(* Logix 5000 project; controller FV vendor 1 type 14 code 217 rev 31.11; software revision 31.00; part 61 of 63 *)
(* tags used below, declared in another part *)
   CWD : CHECKWORD_FLAGS;
   FV_N88 : INT[255];   // YSP COMMS Data transferred to/ from yeast press PLC
   One_Second_One_Scan : ALIAS FOR One_Second_1_scan;
   YP_B103 : INT[15];   // Original N File From SLC, No Description Available
   YP_BLUNG_OV : PlantItem;   // BLUNG_OV
   YP_BLUNG_OV_RawInput : ALIAS FOR RIO_Rack_3:2:I.Data.1;   // YP_BLUNG_OV
   YP_CONV_STOP : PlantItem;   // CONV_STOP
   YP_CONV_STOP_RawInput : ALIAS FOR RIO_Rack_3:2:I.Data.7;   // YP_CONV_STOP
   YP_INP1 : PlantItem;   // INP1
   YP_INP10 : PlantItem;   // INP10
   YP_INP10_RawInput : ALIAS FOR RIO_Rack_3:2:I.Data.14;   // YP_INP10
   YP_INP11 : PlantItem;   // INP11
   YP_INP11_RawInput : ALIAS FOR RIO_Rack_3:2:I.Data.15;   // YP_INP11
   YP_INP1_RawInput : ALIAS FOR RIO_Rack_3:2:I.Data.2;   // YP_INP1
   YP_INP2 : PlantItem;   // INP2
   YP_INP2_RawInput : ALIAS FOR RIO_Rack_3:2:I.Data.3;   // YP_INP2
   YP_INP3 : PlantItem;   // INP3
   YP_INP3_RawInput : ALIAS FOR RIO_Rack_3:2:I.Data.4;   // YP_INP3
   YP_INP4 : PlantItem;   // INP4
   YP_INP4_RawInput : ALIAS FOR RIO_Rack_3:2:I.Data.8;   // YP_INP4
   YP_INP5 : PlantItem;   // INP5
   YP_INP5_RawInput : ALIAS FOR RIO_Rack_3:2:I.Data.9;   // YP_INP5
   YP_INP6 : PlantItem;   // INP6
   YP_INP6_RawInput : ALIAS FOR RIO_Rack_3:2:I.Data.10;   // YP_INP6
   YP_INP7 : PlantItem;   // INP7
   YP_INP7_RawInput : ALIAS FOR RIO_Rack_3:2:I.Data.11;   // YP_INP7
   YP_INP8 : PlantItem;   // INP8
   YP_INP8_RawInput : ALIAS FOR RIO_Rack_3:2:I.Data.12;   // YP_INP8
   YP_INP9 : PlantItem;   // INP9
   YP_INP9_RawInput : ALIAS FOR RIO_Rack_3:2:I.Data.13;   // YP_INP9
   YP_N10 : INT[105];   // COMMS BLOC comms block to fv pl c
   YP_N40 : INT[9];   // Original N File From SLC, No Description Available
   YP_N55 : INT[244];   // Original N File From SLC, No Description Available
   YP_N7 : INT[56];   // INTEGER
   YP_PILZ_OK : PlantItem;   // PILZ_OK
   YP_PILZ_OK_RawInput : ALIAS FOR RIO_Rack_3:2:I.Data.0;   // YP_PILZ_OK
   YP_PRESS_CL : PlantItem;   // PRESS_CL
   YP_PRESS_CL_RawInput : ALIAS FOR RIO_Rack_3:2:I.Data.5;   // YP_PRESS_CL
   YP_PRESS_OP : PlantItem;   // PRESS_OP
   YP_PRESS_OP_RawInput : ALIAS FOR RIO_Rack_3:2:I.Data.6;   // YP_PRESS_OP
   YP_T21 : TIMER[30];
   YP_YST1_HL : PlantItem;   // YST1_HL
   YP_YST1_HL_RawInput : ALIAS FOR RIO_Rack_3:1:I.Data.1;   // YP_YST1_HL
   YP_YST2_HL : PlantItem;   // YST2_HL
   YP_YST2_HL_RawInput : ALIAS FOR RIO_Rack_3:1:I.Data.3;   // YP_YST2_HL
(* YP_Common, continued *)

ROUTINE YP_BLUNGER_14   (* ladder *)
   0: XIO(YP_N40[2].0)XIO(YP_N40[2].1)OTL(YP_N40[2].0);
   1: XIC(YP_N40[2].1)XIO(YP_B103[3].0)[GRT(YP_T21[1].ACC,YP_N55[30]) ,XIC(YP_B103[3].1) ][OTU(YP_N40[2].1) ,OTL(YP_N40[2].0) ];
   2: XIC(YP_N40[2].0)XIC(YP_B103[3].0)[OTU(YP_N40[2].0) ,OTL(YP_N40[2].1) ];
   3: EQU(YP_N55[31],0)MOV(YP_N55[32],YP_N55[30]);
   4: EQU(YP_N55[31],1)MOV(YP_N55[33],YP_N55[30]);
   5: EQU(YP_N55[31],2)MOV(YP_N55[34],YP_N55[30]);
   6: XIC(YP_N40[2].1)TON(YP_T21[1],?,?);
   7: XIO(YP_N40[3].0)XIO(YP_N40[3].1)OTL(YP_N40[3].0);
   8: XIC(YP_N40[3].1)[GRT(YP_T21[2].ACC,YP_N55[40]) ,XIC(YP_B103[3].3) ,XIC(YP_N7[38].0) ,XIC(YP_N7[38].1) ][OTU(YP_N40[3].1) ,OTL(YP_N40[3].0) ];
   9: XIC(YP_N40[3].0)XIC(YP_B103[3].2)[OTU(YP_N40[3].0) ,OTL(YP_N40[3].1) ];
   10: EQU(YP_N55[41],0)MOV(YP_N55[42],YP_N55[40]);
   11: EQU(YP_N55[41],1)MOV(YP_N55[43],YP_N55[40]);
   12: EQU(YP_N55[41],2)MOV(YP_N55[44],YP_N55[40]);
   13: XIC(YP_N40[3].1)TON(YP_T21[2],?,?);
   14: XIC(YP_N40[3].1)XIC(YP_N7[40].0)EQU(YP_N7[39],1)OTL(YP_N7[38].0);
   15: XIC(YP_N40[3].1)XIC(YP_N7[40].1)EQU(YP_N7[39],2)OTL(YP_N7[38].1);
   16: XIC(YP_N40[3].1)EQU(YP_N7[39],99)OTE(YP_N7[38].2);
END_ROUTINE

ROUTINE YP_COMMS_4   (* ladder *)
   0: XIO(YP_T21[3].DN)TON(YP_T21[3],?,?);
   1: XIC(YP_T21[3].DN)COP(FV_N88[0],YP_N10[10],2);
   2: EQU(YP_N10[11],99)MOV(99,YP_N7[39]);
   3: EQU(YP_N10[11],1)MOV(1,YP_N7[39]);
   4: EQU(YP_N10[11],2)MOV(2,YP_N7[39]);
   5: XIC(YP_N7[38].0)OTE(YP_N10[1].0);
   6: XIC(YP_N7[38].1)OTE(YP_N10[1].1);
   7: XIC(YP_N10[10].0)OTE(YP_N10[0].0);
END_ROUTINE

ROUTINE YP_Digital_Inputs   (* ladder *)
   0: [XIC(S:FS) OTU(YP_YST1_HL.CW.[CWD.MANUAL]) ,[XIC(YP_YST1_HL_RawInput) XIO(YP_YST1_HL.CW.[CWD.MANUAL]) ,XIC(YP_YST1_HL.CW.[CWD.MANDRV]) XIC(YP_YST1_HL.CW.[CWD.MANUAL]) ] OTE(YP_YST1_HL.CW.[CWD.INPUTSTATUS]) ,XIC(One_Second_One_Scan) [XIC(YP_YST1_HL.CW.[CWD.INPUTSTATUS]) XIO(YP_YST1_HL.CW.[CWD.INPUTSTATUSDEBOUNCED]) ,XIO(YP_YST1_HL.CW.[CWD.INPUTSTATUS]) XIC(YP_YST1_HL.CW.[CWD.INPUTSTATUSDEBOUNCED]) ] ADD(1,YP_YST1_HL.DebounceTimer,YP_YST1_HL.DebounceTimer) ,[XIC(YP_YST1_HL.CW.[CWD.INPUTSTATUS]) XIC(YP_YST1_HL.CW.[CWD.INPUTSTATUSDEBOUNCED]) ,XIO(YP_YST1_HL.CW.[CWD.INPUTSTATUS]) XIO(YP_YST1_HL.CW.[CWD.INPUTSTATUSDEBOUNCED]) ] CLR(YP_YST1_HL.DebounceTimer) ,GEQ(YP_YST1_HL.DebounceTimer,YP_YST1_HL.DebounceTime) XIC(YP_YST1_HL.CW.[CWD.INPUTSTATUS]) [OTL(YP_YST1_HL.CW.[CWD.INPUTSTATUSDEBOUNCED]) ,CLR(YP_YST1_HL.DebounceTimer) ] ,GEQ(YP_YST1_HL.DebounceTimer,YP_YST1_HL.DebounceTime) XIO(YP_YST1_HL.CW.[CWD.INPUTSTATUS]) [OTU(YP_YST1_HL.CW.[CWD.INPUTSTATUSDEBOUNCED]) ,CLR(YP_YST1_HL.DebounceTimer) ] ];
   1: [XIC(S:FS) OTU(YP_YST2_HL.CW.[CWD.MANUAL]) ,[XIC(YP_YST2_HL_RawInput) XIO(YP_YST2_HL.CW.[CWD.MANUAL]) ,XIC(YP_YST2_HL.CW.[CWD.MANDRV]) XIC(YP_YST2_HL.CW.[CWD.MANUAL]) ] OTE(YP_YST2_HL.CW.[CWD.INPUTSTATUS]) ,XIC(One_Second_One_Scan) [XIC(YP_YST2_HL.CW.[CWD.INPUTSTATUS]) XIO(YP_YST2_HL.CW.[CWD.INPUTSTATUSDEBOUNCED]) ,XIO(YP_YST2_HL.CW.[CWD.INPUTSTATUS]) XIC(YP_YST2_HL.CW.[CWD.INPUTSTATUSDEBOUNCED]) ] ADD(1,YP_YST2_HL.DebounceTimer,YP_YST2_HL.DebounceTimer) ,[XIC(YP_YST2_HL.CW.[CWD.INPUTSTATUS]) XIC(YP_YST2_HL.CW.[CWD.INPUTSTATUSDEBOUNCED]) ,XIO(YP_YST2_HL.CW.[CWD.INPUTSTATUS]) XIO(YP_YST2_HL.CW.[CWD.INPUTSTATUSDEBOUNCED]) ] CLR(YP_YST2_HL.DebounceTimer) ,GEQ(YP_YST2_HL.DebounceTimer,YP_YST2_HL.DebounceTime) XIC(YP_YST2_HL.CW.[CWD.INPUTSTATUS]) [OTL(YP_YST2_HL.CW.[CWD.INPUTSTATUSDEBOUNCED]) ,CLR(YP_YST2_HL.DebounceTimer) ] ,GEQ(YP_YST2_HL.DebounceTimer,YP_YST2_HL.DebounceTime) XIO(YP_YST2_HL.CW.[CWD.INPUTSTATUS]) [OTU(YP_YST2_HL.CW.[CWD.INPUTSTATUSDEBOUNCED]) ,CLR(YP_YST2_HL.DebounceTimer) ] ];
   2: [XIC(S:FS) OTU(YP_PILZ_OK.CW.[CWD.MANUAL]) ,[XIC(YP_PILZ_OK_RawInput) XIO(YP_PILZ_OK.CW.[CWD.MANUAL]) ,XIC(YP_PILZ_OK.CW.[CWD.MANDRV]) XIC(YP_PILZ_OK.CW.[CWD.MANUAL]) ] OTE(YP_PILZ_OK.CW.[CWD.INPUTSTATUS]) ,XIC(One_Second_One_Scan) [XIC(YP_PILZ_OK.CW.[CWD.INPUTSTATUS]) XIO(YP_PILZ_OK.CW.[CWD.INPUTSTATUSDEBOUNCED]) ,XIO(YP_PILZ_OK.CW.[CWD.INPUTSTATUS]) XIC(YP_PILZ_OK.CW.[CWD.INPUTSTATUSDEBOUNCED]) ] ADD(1,YP_PILZ_OK.DebounceTimer,YP_PILZ_OK.DebounceTimer) ,[XIC(YP_PILZ_OK.CW.[CWD.INPUTSTATUS]) XIC(YP_PILZ_OK.CW.[CWD.INPUTSTATUSDEBOUNCED]) ,XIO(YP_PILZ_OK.CW.[CWD.INPUTSTATUS]) XIO(YP_PILZ_OK.CW.[CWD.INPUTSTATUSDEBOUNCED]) ] CLR(YP_PILZ_OK.DebounceTimer) ,GEQ(YP_PILZ_OK.DebounceTimer,YP_PILZ_OK.DebounceTime) XIC(YP_PILZ_OK.CW.[CWD.INPUTSTATUS]) [OTL(YP_PILZ_OK.CW.[CWD.INPUTSTATUSDEBOUNCED]) ,CLR(YP_PILZ_OK.DebounceTimer) ] ,GEQ(YP_PILZ_OK.DebounceTimer,YP_PILZ_OK.DebounceTime) XIO(YP_PILZ_OK.CW.[CWD.INPUTSTATUS]) [OTU(YP_PILZ_OK.CW.[CWD.INPUTSTATUSDEBOUNCED]) ,CLR(YP_PILZ_OK.DebounceTimer) ] ];
   3: [XIC(S:FS) OTU(YP_BLUNG_OV.CW.[CWD.MANUAL]) ,[XIC(YP_BLUNG_OV_RawInput) XIO(YP_BLUNG_OV.CW.[CWD.MANUAL]) ,XIC(YP_BLUNG_OV.CW.[CWD.MANDRV]) XIC(YP_BLUNG_OV.CW.[CWD.MANUAL]) ] OTE(YP_BLUNG_OV.CW.[CWD.INPUTSTATUS]) ,XIC(One_Second_One_Scan) [XIC(YP_BLUNG_OV.CW.[CWD.INPUTSTATUS]) XIO(YP_BLUNG_OV.CW.[CWD.INPUTSTATUSDEBOUNCED]) ,XIO(YP_BLUNG_OV.CW.[CWD.INPUTSTATUS]) XIC(YP_BLUNG_OV.CW.[CWD.INPUTSTATUSDEBOUNCED]) ] ADD(1,YP_BLUNG_OV.DebounceTimer,YP_BLUNG_OV.DebounceTimer) ,[XIC(YP_BLUNG_OV.CW.[CWD.INPUTSTATUS]) XIC(YP_BLUNG_OV.CW.[CWD.INPUTSTATUSDEBOUNCED]) ,XIO(YP_BLUNG_OV.CW.[CWD.INPUTSTATUS]) XIO(YP_BLUNG_OV.CW.[CWD.INPUTSTATUSDEBOUNCED]) ] CLR(YP_BLUNG_OV.DebounceTimer) ,GEQ(YP_BLUNG_OV.DebounceTimer,YP_BLUNG_OV.DebounceTime) XIC(YP_BLUNG_OV.CW.[CWD.INPUTSTATUS]) [OTL(YP_BLUNG_OV.CW.[CWD.INPUTSTATUSDEBOUNCED]) ,CLR(YP_BLUNG_OV.DebounceTimer) ] ,GEQ(YP_BLUNG_OV.DebounceTimer,YP_BLUNG_OV.DebounceTime) XIO(YP_BLUNG_OV.CW.[CWD.INPUTSTATUS]) [OTU(YP_BLUNG_OV.CW.[CWD.INPUTSTATUSDEBOUNCED]) ,CLR(YP_BLUNG_OV.DebounceTimer) ] ];
   4: [XIC(S:FS) OTU(YP_INP1.CW.[CWD.MANUAL]) ,[XIC(YP_INP1_RawInput) XIO(YP_INP1.CW.[CWD.MANUAL]) ,XIC(YP_INP1.CW.[CWD.MANDRV]) XIC(YP_INP1.CW.[CWD.MANUAL]) ] OTE(YP_INP1.CW.[CWD.INPUTSTATUS]) ,XIC(One_Second_One_Scan) [XIC(YP_INP1.CW.[CWD.INPUTSTATUS]) XIO(YP_INP1.CW.[CWD.INPUTSTATUSDEBOUNCED]) ,XIO(YP_INP1.CW.[CWD.INPUTSTATUS]) XIC(YP_INP1.CW.[CWD.INPUTSTATUSDEBOUNCED]) ] ADD(1,YP_INP1.DebounceTimer,YP_INP1.DebounceTimer) ,[XIC(YP_INP1.CW.[CWD.INPUTSTATUS]) XIC(YP_INP1.CW.[CWD.INPUTSTATUSDEBOUNCED]) ,XIO(YP_INP1.CW.[CWD.INPUTSTATUS]) XIO(YP_INP1.CW.[CWD.INPUTSTATUSDEBOUNCED]) ] CLR(YP_INP1.DebounceTimer) ,GEQ(YP_INP1.DebounceTimer,YP_INP1.DebounceTime) XIC(YP_INP1.CW.[CWD.INPUTSTATUS]) [OTL(YP_INP1.CW.[CWD.INPUTSTATUSDEBOUNCED]) ,CLR(YP_INP1.DebounceTimer) ] ,GEQ(YP_INP1.DebounceTimer,YP_INP1.DebounceTime) XIO(YP_INP1.CW.[CWD.INPUTSTATUS]) [OTU(YP_INP1.CW.[CWD.INPUTSTATUSDEBOUNCED]) ,CLR(YP_INP1.DebounceTimer) ] ];
   5: [XIC(S:FS) OTU(YP_INP2.CW.[CWD.MANUAL]) ,[XIC(YP_INP2_RawInput) XIO(YP_INP2.CW.[CWD.MANUAL]) ,XIC(YP_INP2.CW.[CWD.MANDRV]) XIC(YP_INP2.CW.[CWD.MANUAL]) ] OTE(YP_INP2.CW.[CWD.INPUTSTATUS]) ,XIC(One_Second_One_Scan) [XIC(YP_INP2.CW.[CWD.INPUTSTATUS]) XIO(YP_INP2.CW.[CWD.INPUTSTATUSDEBOUNCED]) ,XIO(YP_INP2.CW.[CWD.INPUTSTATUS]) XIC(YP_INP2.CW.[CWD.INPUTSTATUSDEBOUNCED]) ] ADD(1,YP_INP2.DebounceTimer,YP_INP2.DebounceTimer) ,[XIC(YP_INP2.CW.[CWD.INPUTSTATUS]) XIC(YP_INP2.CW.[CWD.INPUTSTATUSDEBOUNCED]) ,XIO(YP_INP2.CW.[CWD.INPUTSTATUS]) XIO(YP_INP2.CW.[CWD.INPUTSTATUSDEBOUNCED]) ] CLR(YP_INP2.DebounceTimer) ,GEQ(YP_INP2.DebounceTimer,YP_INP2.DebounceTime) XIC(YP_INP2.CW.[CWD.INPUTSTATUS]) [OTL(YP_INP2.CW.[CWD.INPUTSTATUSDEBOUNCED]) ,CLR(YP_INP2.DebounceTimer) ] ,GEQ(YP_INP2.DebounceTimer,YP_INP2.DebounceTime) XIO(YP_INP2.CW.[CWD.INPUTSTATUS]) [OTU(YP_INP2.CW.[CWD.INPUTSTATUSDEBOUNCED]) ,CLR(YP_INP2.DebounceTimer) ] ];
   6: [XIC(S:FS) OTU(YP_INP3.CW.[CWD.MANUAL]) ,[XIC(YP_INP3_RawInput) XIO(YP_INP3.CW.[CWD.MANUAL]) ,XIC(YP_INP3.CW.[CWD.MANDRV]) XIC(YP_INP3.CW.[CWD.MANUAL]) ] OTE(YP_INP3.CW.[CWD.INPUTSTATUS]) ,XIC(One_Second_One_Scan) [XIC(YP_INP3.CW.[CWD.INPUTSTATUS]) XIO(YP_INP3.CW.[CWD.INPUTSTATUSDEBOUNCED]) ,XIO(YP_INP3.CW.[CWD.INPUTSTATUS]) XIC(YP_INP3.CW.[CWD.INPUTSTATUSDEBOUNCED]) ] ADD(1,YP_INP3.DebounceTimer,YP_INP3.DebounceTimer) ,[XIC(YP_INP3.CW.[CWD.INPUTSTATUS]) XIC(YP_INP3.CW.[CWD.INPUTSTATUSDEBOUNCED]) ,XIO(YP_INP3.CW.[CWD.INPUTSTATUS]) XIO(YP_INP3.CW.[CWD.INPUTSTATUSDEBOUNCED]) ] CLR(YP_INP3.DebounceTimer) ,GEQ(YP_INP3.DebounceTimer,YP_INP3.DebounceTime) XIC(YP_INP3.CW.[CWD.INPUTSTATUS]) [OTL(YP_INP3.CW.[CWD.INPUTSTATUSDEBOUNCED]) ,CLR(YP_INP3.DebounceTimer) ] ,GEQ(YP_INP3.DebounceTimer,YP_INP3.DebounceTime) XIO(YP_INP3.CW.[CWD.INPUTSTATUS]) [OTU(YP_INP3.CW.[CWD.INPUTSTATUSDEBOUNCED]) ,CLR(YP_INP3.DebounceTimer) ] ];
   7: [XIC(S:FS) OTU(YP_PRESS_CL.CW.[CWD.MANUAL]) ,[XIC(YP_PRESS_CL_RawInput) XIO(YP_PRESS_CL.CW.[CWD.MANUAL]) ,XIC(YP_PRESS_CL.CW.[CWD.MANDRV]) XIC(YP_PRESS_CL.CW.[CWD.MANUAL]) ] OTE(YP_PRESS_CL.CW.[CWD.INPUTSTATUS]) ,XIC(One_Second_One_Scan) [XIC(YP_PRESS_CL.CW.[CWD.INPUTSTATUS]) XIO(YP_PRESS_CL.CW.[CWD.INPUTSTATUSDEBOUNCED]) ,XIO(YP_PRESS_CL.CW.[CWD.INPUTSTATUS]) XIC(YP_PRESS_CL.CW.[CWD.INPUTSTATUSDEBOUNCED]) ] ADD(1,YP_PRESS_CL.DebounceTimer,YP_PRESS_CL.DebounceTimer) ,[XIC(YP_PRESS_CL.CW.[CWD.INPUTSTATUS]) XIC(YP_PRESS_CL.CW.[CWD.INPUTSTATUSDEBOUNCED]) ,XIO(YP_PRESS_CL.CW.[CWD.INPUTSTATUS]) XIO(YP_PRESS_CL.CW.[CWD.INPUTSTATUSDEBOUNCED]) ] CLR(YP_PRESS_CL.DebounceTimer) ,GEQ(YP_PRESS_CL.DebounceTimer,YP_PRESS_CL.DebounceTime) XIC(YP_PRESS_CL.CW.[CWD.INPUTSTATUS]) [OTL(YP_PRESS_CL.CW.[CWD.INPUTSTATUSDEBOUNCED]) ,CLR(YP_PRESS_CL.DebounceTimer) ] ,GEQ(YP_PRESS_CL.DebounceTimer,YP_PRESS_CL.DebounceTime) XIO(YP_PRESS_CL.CW.[CWD.INPUTSTATUS]) [OTU(YP_PRESS_CL.CW.[CWD.INPUTSTATUSDEBOUNCED]) ,CLR(YP_PRESS_CL.DebounceTimer) ] ];
   8: [XIC(S:FS) OTU(YP_PRESS_OP.CW.[CWD.MANUAL]) ,[XIC(YP_PRESS_OP_RawInput) XIO(YP_PRESS_OP.CW.[CWD.MANUAL]) ,XIC(YP_PRESS_OP.CW.[CWD.MANDRV]) XIC(YP_PRESS_OP.CW.[CWD.MANUAL]) ] OTE(YP_PRESS_OP.CW.[CWD.INPUTSTATUS]) ,XIC(One_Second_One_Scan) [XIC(YP_PRESS_OP.CW.[CWD.INPUTSTATUS]) XIO(YP_PRESS_OP.CW.[CWD.INPUTSTATUSDEBOUNCED]) ,XIO(YP_PRESS_OP.CW.[CWD.INPUTSTATUS]) XIC(YP_PRESS_OP.CW.[CWD.INPUTSTATUSDEBOUNCED]) ] ADD(1,YP_PRESS_OP.DebounceTimer,YP_PRESS_OP.DebounceTimer) ,[XIC(YP_PRESS_OP.CW.[CWD.INPUTSTATUS]) XIC(YP_PRESS_OP.CW.[CWD.INPUTSTATUSDEBOUNCED]) ,XIO(YP_PRESS_OP.CW.[CWD.INPUTSTATUS]) XIO(YP_PRESS_OP.CW.[CWD.INPUTSTATUSDEBOUNCED]) ] CLR(YP_PRESS_OP.DebounceTimer) ,GEQ(YP_PRESS_OP.DebounceTimer,YP_PRESS_OP.DebounceTime) XIC(YP_PRESS_OP.CW.[CWD.INPUTSTATUS]) [OTL(YP_PRESS_OP.CW.[CWD.INPUTSTATUSDEBOUNCED]) ,CLR(YP_PRESS_OP.DebounceTimer) ] ,GEQ(YP_PRESS_OP.DebounceTimer,YP_PRESS_OP.DebounceTime) XIO(YP_PRESS_OP.CW.[CWD.INPUTSTATUS]) [OTU(YP_PRESS_OP.CW.[CWD.INPUTSTATUSDEBOUNCED]) ,CLR(YP_PRESS_OP.DebounceTimer) ] ];
   9: [XIC(S:FS) OTU(YP_CONV_STOP.CW.[CWD.MANUAL]) ,[XIC(YP_CONV_STOP_RawInput) XIO(YP_CONV_STOP.CW.[CWD.MANUAL]) ,XIC(YP_CONV_STOP.CW.[CWD.MANDRV]) XIC(YP_CONV_STOP.CW.[CWD.MANUAL]) ] OTE(YP_CONV_STOP.CW.[CWD.INPUTSTATUS]) ,XIC(One_Second_One_Scan) [XIC(YP_CONV_STOP.CW.[CWD.INPUTSTATUS]) XIO(YP_CONV_STOP.CW.[CWD.INPUTSTATUSDEBOUNCED]) ,XIO(YP_CONV_STOP.CW.[CWD.INPUTSTATUS]) XIC(YP_CONV_STOP.CW.[CWD.INPUTSTATUSDEBOUNCED]) ] ADD(1,YP_CONV_STOP.DebounceTimer,YP_CONV_STOP.DebounceTimer) ,[XIC(YP_CONV_STOP.CW.[CWD.INPUTSTATUS]) XIC(YP_CONV_STOP.CW.[CWD.INPUTSTATUSDEBOUNCED]) ,XIO(YP_CONV_STOP.CW.[CWD.INPUTSTATUS]) XIO(YP_CONV_STOP.CW.[CWD.INPUTSTATUSDEBOUNCED]) ] CLR(YP_CONV_STOP.DebounceTimer) ,GEQ(YP_CONV_STOP.DebounceTimer,YP_CONV_STOP.DebounceTime) XIC(YP_CONV_STOP.CW.[CWD.INPUTSTATUS]) [OTL(YP_CONV_STOP.CW.[CWD.INPUTSTATUSDEBOUNCED]) ,CLR(YP_CONV_STOP.DebounceTimer) ] ,GEQ(YP_CONV_STOP.DebounceTimer,YP_CONV_STOP.DebounceTime) XIO(YP_CONV_STOP.CW.[CWD.INPUTSTATUS]) [OTU(YP_CONV_STOP.CW.[CWD.INPUTSTATUSDEBOUNCED]) ,CLR(YP_CONV_STOP.DebounceTimer) ] ];
   10: [XIC(S:FS) OTU(YP_INP4.CW.[CWD.MANUAL]) ,[XIC(YP_INP4_RawInput) XIO(YP_INP4.CW.[CWD.MANUAL]) ,XIC(YP_INP4.CW.[CWD.MANDRV]) XIC(YP_INP4.CW.[CWD.MANUAL]) ] OTE(YP_INP4.CW.[CWD.INPUTSTATUS]) ,XIC(One_Second_One_Scan) [XIC(YP_INP4.CW.[CWD.INPUTSTATUS]) XIO(YP_INP4.CW.[CWD.INPUTSTATUSDEBOUNCED]) ,XIO(YP_INP4.CW.[CWD.INPUTSTATUS]) XIC(YP_INP4.CW.[CWD.INPUTSTATUSDEBOUNCED]) ] ADD(1,YP_INP4.DebounceTimer,YP_INP4.DebounceTimer) ,[XIC(YP_INP4.CW.[CWD.INPUTSTATUS]) XIC(YP_INP4.CW.[CWD.INPUTSTATUSDEBOUNCED]) ,XIO(YP_INP4.CW.[CWD.INPUTSTATUS]) XIO(YP_INP4.CW.[CWD.INPUTSTATUSDEBOUNCED]) ] CLR(YP_INP4.DebounceTimer) ,GEQ(YP_INP4.DebounceTimer,YP_INP4.DebounceTime) XIC(YP_INP4.CW.[CWD.INPUTSTATUS]) [OTL(YP_INP4.CW.[CWD.INPUTSTATUSDEBOUNCED]) ,CLR(YP_INP4.DebounceTimer) ] ,GEQ(YP_INP4.DebounceTimer,YP_INP4.DebounceTime) XIO(YP_INP4.CW.[CWD.INPUTSTATUS]) [OTU(YP_INP4.CW.[CWD.INPUTSTATUSDEBOUNCED]) ,CLR(YP_INP4.DebounceTimer) ] ];
   11: [XIC(S:FS) OTU(YP_INP5.CW.[CWD.MANUAL]) ,[XIC(YP_INP5_RawInput) XIO(YP_INP5.CW.[CWD.MANUAL]) ,XIC(YP_INP5.CW.[CWD.MANDRV]) XIC(YP_INP5.CW.[CWD.MANUAL]) ] OTE(YP_INP5.CW.[CWD.INPUTSTATUS]) ,XIC(One_Second_One_Scan) [XIC(YP_INP5.CW.[CWD.INPUTSTATUS]) XIO(YP_INP5.CW.[CWD.INPUTSTATUSDEBOUNCED]) ,XIO(YP_INP5.CW.[CWD.INPUTSTATUS]) XIC(YP_INP5.CW.[CWD.INPUTSTATUSDEBOUNCED]) ] ADD(1,YP_INP5.DebounceTimer,YP_INP5.DebounceTimer) ,[XIC(YP_INP5.CW.[CWD.INPUTSTATUS]) XIC(YP_INP5.CW.[CWD.INPUTSTATUSDEBOUNCED]) ,XIO(YP_INP5.CW.[CWD.INPUTSTATUS]) XIO(YP_INP5.CW.[CWD.INPUTSTATUSDEBOUNCED]) ] CLR(YP_INP5.DebounceTimer) ,GEQ(YP_INP5.DebounceTimer,YP_INP5.DebounceTime) XIC(YP_INP5.CW.[CWD.INPUTSTATUS]) [OTL(YP_INP5.CW.[CWD.INPUTSTATUSDEBOUNCED]) ,CLR(YP_INP5.DebounceTimer) ] ,GEQ(YP_INP5.DebounceTimer,YP_INP5.DebounceTime) XIO(YP_INP5.CW.[CWD.INPUTSTATUS]) [OTU(YP_INP5.CW.[CWD.INPUTSTATUSDEBOUNCED]) ,CLR(YP_INP5.DebounceTimer) ] ];
   12: [XIC(S:FS) OTU(YP_INP6.CW.[CWD.MANUAL]) ,[XIC(YP_INP6_RawInput) XIO(YP_INP6.CW.[CWD.MANUAL]) ,XIC(YP_INP6.CW.[CWD.MANDRV]) XIC(YP_INP6.CW.[CWD.MANUAL]) ] OTE(YP_INP6.CW.[CWD.INPUTSTATUS]) ,XIC(One_Second_One_Scan) [XIC(YP_INP6.CW.[CWD.INPUTSTATUS]) XIO(YP_INP6.CW.[CWD.INPUTSTATUSDEBOUNCED]) ,XIO(YP_INP6.CW.[CWD.INPUTSTATUS]) XIC(YP_INP6.CW.[CWD.INPUTSTATUSDEBOUNCED]) ] ADD(1,YP_INP6.DebounceTimer,YP_INP6.DebounceTimer) ,[XIC(YP_INP6.CW.[CWD.INPUTSTATUS]) XIC(YP_INP6.CW.[CWD.INPUTSTATUSDEBOUNCED]) ,XIO(YP_INP6.CW.[CWD.INPUTSTATUS]) XIO(YP_INP6.CW.[CWD.INPUTSTATUSDEBOUNCED]) ] CLR(YP_INP6.DebounceTimer) ,GEQ(YP_INP6.DebounceTimer,YP_INP6.DebounceTime) XIC(YP_INP6.CW.[CWD.INPUTSTATUS]) [OTL(YP_INP6.CW.[CWD.INPUTSTATUSDEBOUNCED]) ,CLR(YP_INP6.DebounceTimer) ] ,GEQ(YP_INP6.DebounceTimer,YP_INP6.DebounceTime) XIO(YP_INP6.CW.[CWD.INPUTSTATUS]) [OTU(YP_INP6.CW.[CWD.INPUTSTATUSDEBOUNCED]) ,CLR(YP_INP6.DebounceTimer) ] ];
   13: [XIC(S:FS) OTU(YP_INP7.CW.[CWD.MANUAL]) ,[XIC(YP_INP7_RawInput) XIO(YP_INP7.CW.[CWD.MANUAL]) ,XIC(YP_INP7.CW.[CWD.MANDRV]) XIC(YP_INP7.CW.[CWD.MANUAL]) ] OTE(YP_INP7.CW.[CWD.INPUTSTATUS]) ,XIC(One_Second_One_Scan) [XIC(YP_INP7.CW.[CWD.INPUTSTATUS]) XIO(YP_INP7.CW.[CWD.INPUTSTATUSDEBOUNCED]) ,XIO(YP_INP7.CW.[CWD.INPUTSTATUS]) XIC(YP_INP7.CW.[CWD.INPUTSTATUSDEBOUNCED]) ] ADD(1,YP_INP7.DebounceTimer,YP_INP7.DebounceTimer) ,[XIC(YP_INP7.CW.[CWD.INPUTSTATUS]) XIC(YP_INP7.CW.[CWD.INPUTSTATUSDEBOUNCED]) ,XIO(YP_INP7.CW.[CWD.INPUTSTATUS]) XIO(YP_INP7.CW.[CWD.INPUTSTATUSDEBOUNCED]) ] CLR(YP_INP7.DebounceTimer) ,GEQ(YP_INP7.DebounceTimer,YP_INP7.DebounceTime) XIC(YP_INP7.CW.[CWD.INPUTSTATUS]) [OTL(YP_INP7.CW.[CWD.INPUTSTATUSDEBOUNCED]) ,CLR(YP_INP7.DebounceTimer) ] ,GEQ(YP_INP7.DebounceTimer,YP_INP7.DebounceTime) XIO(YP_INP7.CW.[CWD.INPUTSTATUS]) [OTU(YP_INP7.CW.[CWD.INPUTSTATUSDEBOUNCED]) ,CLR(YP_INP7.DebounceTimer) ] ];
   14: [XIC(S:FS) OTU(YP_INP8.CW.[CWD.MANUAL]) ,[XIC(YP_INP8_RawInput) XIO(YP_INP8.CW.[CWD.MANUAL]) ,XIC(YP_INP8.CW.[CWD.MANDRV]) XIC(YP_INP8.CW.[CWD.MANUAL]) ] OTE(YP_INP8.CW.[CWD.INPUTSTATUS]) ,XIC(One_Second_One_Scan) [XIC(YP_INP8.CW.[CWD.INPUTSTATUS]) XIO(YP_INP8.CW.[CWD.INPUTSTATUSDEBOUNCED]) ,XIO(YP_INP8.CW.[CWD.INPUTSTATUS]) XIC(YP_INP8.CW.[CWD.INPUTSTATUSDEBOUNCED]) ] ADD(1,YP_INP8.DebounceTimer,YP_INP8.DebounceTimer) ,[XIC(YP_INP8.CW.[CWD.INPUTSTATUS]) XIC(YP_INP8.CW.[CWD.INPUTSTATUSDEBOUNCED]) ,XIO(YP_INP8.CW.[CWD.INPUTSTATUS]) XIO(YP_INP8.CW.[CWD.INPUTSTATUSDEBOUNCED]) ] CLR(YP_INP8.DebounceTimer) ,GEQ(YP_INP8.DebounceTimer,YP_INP8.DebounceTime) XIC(YP_INP8.CW.[CWD.INPUTSTATUS]) [OTL(YP_INP8.CW.[CWD.INPUTSTATUSDEBOUNCED]) ,CLR(YP_INP8.DebounceTimer) ] ,GEQ(YP_INP8.DebounceTimer,YP_INP8.DebounceTime) XIO(YP_INP8.CW.[CWD.INPUTSTATUS]) [OTU(YP_INP8.CW.[CWD.INPUTSTATUSDEBOUNCED]) ,CLR(YP_INP8.DebounceTimer) ] ];
   15: [XIC(S:FS) OTU(YP_INP9.CW.[CWD.MANUAL]) ,[XIC(YP_INP9_RawInput) XIO(YP_INP9.CW.[CWD.MANUAL]) ,XIC(YP_INP9.CW.[CWD.MANDRV]) XIC(YP_INP9.CW.[CWD.MANUAL]) ] OTE(YP_INP9.CW.[CWD.INPUTSTATUS]) ,XIC(One_Second_One_Scan) [XIC(YP_INP9.CW.[CWD.INPUTSTATUS]) XIO(YP_INP9.CW.[CWD.INPUTSTATUSDEBOUNCED]) ,XIO(YP_INP9.CW.[CWD.INPUTSTATUS]) XIC(YP_INP9.CW.[CWD.INPUTSTATUSDEBOUNCED]) ] ADD(1,YP_INP9.DebounceTimer,YP_INP9.DebounceTimer) ,[XIC(YP_INP9.CW.[CWD.INPUTSTATUS]) XIC(YP_INP9.CW.[CWD.INPUTSTATUSDEBOUNCED]) ,XIO(YP_INP9.CW.[CWD.INPUTSTATUS]) XIO(YP_INP9.CW.[CWD.INPUTSTATUSDEBOUNCED]) ] CLR(YP_INP9.DebounceTimer) ,GEQ(YP_INP9.DebounceTimer,YP_INP9.DebounceTime) XIC(YP_INP9.CW.[CWD.INPUTSTATUS]) [OTL(YP_INP9.CW.[CWD.INPUTSTATUSDEBOUNCED]) ,CLR(YP_INP9.DebounceTimer) ] ,GEQ(YP_INP9.DebounceTimer,YP_INP9.DebounceTime) XIO(YP_INP9.CW.[CWD.INPUTSTATUS]) [OTU(YP_INP9.CW.[CWD.INPUTSTATUSDEBOUNCED]) ,CLR(YP_INP9.DebounceTimer) ] ];
   16: [XIC(S:FS) OTU(YP_INP10.CW.[CWD.MANUAL]) ,[XIC(YP_INP10_RawInput) XIO(YP_INP10.CW.[CWD.MANUAL]) ,XIC(YP_INP10.CW.[CWD.MANDRV]) XIC(YP_INP10.CW.[CWD.MANUAL]) ] OTE(YP_INP10.CW.[CWD.INPUTSTATUS]) ,XIC(One_Second_One_Scan) [XIC(YP_INP10.CW.[CWD.INPUTSTATUS]) XIO(YP_INP10.CW.[CWD.INPUTSTATUSDEBOUNCED]) ,XIO(YP_INP10.CW.[CWD.INPUTSTATUS]) XIC(YP_INP10.CW.[CWD.INPUTSTATUSDEBOUNCED]) ] ADD(1,YP_INP10.DebounceTimer,YP_INP10.DebounceTimer) ,[XIC(YP_INP10.CW.[CWD.INPUTSTATUS]) XIC(YP_INP10.CW.[CWD.INPUTSTATUSDEBOUNCED]) ,XIO(YP_INP10.CW.[CWD.INPUTSTATUS]) XIO(YP_INP10.CW.[CWD.INPUTSTATUSDEBOUNCED]) ] CLR(YP_INP10.DebounceTimer) ,GEQ(YP_INP10.DebounceTimer,YP_INP10.DebounceTime) XIC(YP_INP10.CW.[CWD.INPUTSTATUS]) [OTL(YP_INP10.CW.[CWD.INPUTSTATUSDEBOUNCED]) ,CLR(YP_INP10.DebounceTimer) ] ,GEQ(YP_INP10.DebounceTimer,YP_INP10.DebounceTime) XIO(YP_INP10.CW.[CWD.INPUTSTATUS]) [OTU(YP_INP10.CW.[CWD.INPUTSTATUSDEBOUNCED]) ,CLR(YP_INP10.DebounceTimer) ] ];
   17: [XIC(S:FS) OTU(YP_INP11.CW.[CWD.MANUAL]) ,[XIC(YP_INP11_RawInput) XIO(YP_INP11.CW.[CWD.MANUAL]) ,XIC(YP_INP11.CW.[CWD.MANDRV]) XIC(YP_INP11.CW.[CWD.MANUAL]) ] OTE(YP_INP11.CW.[CWD.INPUTSTATUS]) ,XIC(One_Second_One_Scan) [XIC(YP_INP11.CW.[CWD.INPUTSTATUS]) XIO(YP_INP11.CW.[CWD.INPUTSTATUSDEBOUNCED]) ,XIO(YP_INP11.CW.[CWD.INPUTSTATUS]) XIC(YP_INP11.CW.[CWD.INPUTSTATUSDEBOUNCED]) ] ADD(1,YP_INP11.DebounceTimer,YP_INP11.DebounceTimer) ,[XIC(YP_INP11.CW.[CWD.INPUTSTATUS]) XIC(YP_INP11.CW.[CWD.INPUTSTATUSDEBOUNCED]) ,XIO(YP_INP11.CW.[CWD.INPUTSTATUS]) XIO(YP_INP11.CW.[CWD.INPUTSTATUSDEBOUNCED]) ] CLR(YP_INP11.DebounceTimer) ,GEQ(YP_INP11.DebounceTimer,YP_INP11.DebounceTime) XIC(YP_INP11.CW.[CWD.INPUTSTATUS]) [OTL(YP_INP11.CW.[CWD.INPUTSTATUSDEBOUNCED]) ,CLR(YP_INP11.DebounceTimer) ] ,GEQ(YP_INP11.DebounceTimer,YP_INP11.DebounceTime) XIO(YP_INP11.CW.[CWD.INPUTSTATUS]) [OTU(YP_INP11.CW.[CWD.INPUTSTATUSDEBOUNCED]) ,CLR(YP_INP11.DebounceTimer) ] ];
END_ROUTINE
